// TIA Portal project "TestEssProtoFreia" (V13) (continued)

         L     #ET_MAX;
         ITD;
         DTR;
         L     #ET_MIN;
         ITD;
         DTR;
         -R;
         T     #INTER_3;  //ETENDUE DE MESURE MAXI - MINI

         L     #VAL_MINI;
         T     #INTER_4;  //ECHELLE MINI

         L     #INTER_1;
         L     #INTER_2;
         *R;
         L     #INTER_3;
         /R;
         L     #INTER_4;
         +R;
         T     #PV;
         JU    NEXT;
END_REGION

REGION Network 3 (STL): Input type : PT100 en °C
   // Input type : PT100 en °C

   C2:   L     #INPUT;
         ITD;
         DTR;
         L     10.0;
         /R;
         T     #INTER_1;



         L     #INTER_1;
         T     #PV;

         JU    NEXT;
END_REGION

REGION Network 4 (STL): Input type : PT100 en K
   // Input type  : PT100 en K

   C3:   L     #INPUT;
         ITD;
         DTR;
         L     10.0;
         /R;
         L     273.0;
         +R;
         T     #INTER_1;



         L     #INTER_1;
         T     #PV;

         JU    NEXT;
END_REGION

REGION Network 5 (STL): Depassement haut de la valeur convertie
   // Dépassement haut et bas process de la valeur
   NEXT: L     #PV;
         L     #PV_SEUILH;  //Test la valeur maximum pour le dépassement haut
         >R;
         =     #ALM_HIGH;

         L     #PV;
         L     #PV_SEUILB;  //Test la valeur minimum pour le dépassement bas
         <R;
         =     #ALM_LOW;
END_REGION

REGION Network 6 (STL): Depassement bas de la valeur convertie
   // Défaut capteur

         L     #INPUT;
         L     #ET_MAX;
         >I;
         O(;
         L     #INPUT;
         L     #ET_MIN;
         <I;
         );
         =     #ALM_TEMP;

         A     #ALM_TEMP;
         S     #ALM_SENSOR;

         AN    #ALM_TEMP;
         A     #ACQ;
         R     #ALM_SENSOR;

         NOP   0;
END_REGION

REGION Network 7 (STL): Recopie des mini et maxi de la mesure
   // Recopie des mini et maxi de la mesure
         L     #VAL_MAXI;  //Charge le maxi
         T     #PV_HIGH;

         L     #VAL_MINI;  //Charge le mini
         T     #PV_LOW;
END_REGION

REGION Network 8 (STL): Gestion du mot de défaut
   // Gestion du mot de défaut
         A     #ALM_SENSOR;
         JCN   High;  //Retourne un défaut capteur dans le mot
         L     3;  //Usually 3
         T     #ANIM;
         JU    Saut;
   High: A     #ALM_HIGH;
         JCN   Low;  //Retourne un dépassement haut dans le mot
         L     2;
         T     #ANIM;
         JU    Saut;
   Low:  A     #ALM_LOW;
         JCN   Fin;  //Retourne un dépassement bas dans le mot
         L     1;  //Usually 3
         T     #ANIM;
         JU    Saut;

   Fin:  L     0;  //Aucun défaut sur la mesure
         T     #ANIM;
   Saut: NOP   0;
END_REGION

REGION Network 9 (STL): Fin du traitement
   // Fin du traitement
   End:  NOP   0;
END_REGION
END_FUNCTION

FUNCTION "CONVERSION R/T" : Void   // FC20, SCL
{ S7_Optimized_Access := 'FALSE' }
VERSION : 0.1
BEGIN

   //#TEMPERATURE_KELVIN := REAL#29.377125832 + (REAL#2.3156100732 * #"RESISTANCE _OHMS") + (REAL#1.2102319168 * 10 ** -03 * SQR(#"RESISTANCE _OHMS"));
   #TEMPERATURE_KELVIN := REAL#29.37713 + (REAL#2.315610 * #"RESISTANCE _OHMS") + (REAL#1.210232 * 10 ** -03 * SQR(#"RESISTANCE _OHMS"));
END_FUNCTION

FUNCTION "Send_to_Epics" : Void   // FC30, LAD
{ S7_Optimized_Access := 'FALSE' }
VERSION : 0.1
   VAR_TEMP   // added for the SCL form of the ladder/FBD networks
      _w1 : Bool;
   END_VAR
BEGIN

REGION Network 1 (STL): Send timer
         AN    "EPICS_send_T1";
         L     s5t#100ms;
         SD    "EPICS_send_T0";
         A     "EPICS_send_T0";
         L     s5t#100ms;
         SD    "EPICS_send_T1";
         =     "EPICS_do_send";
END_REGION

REGION Network 2: Set ACT_SEND
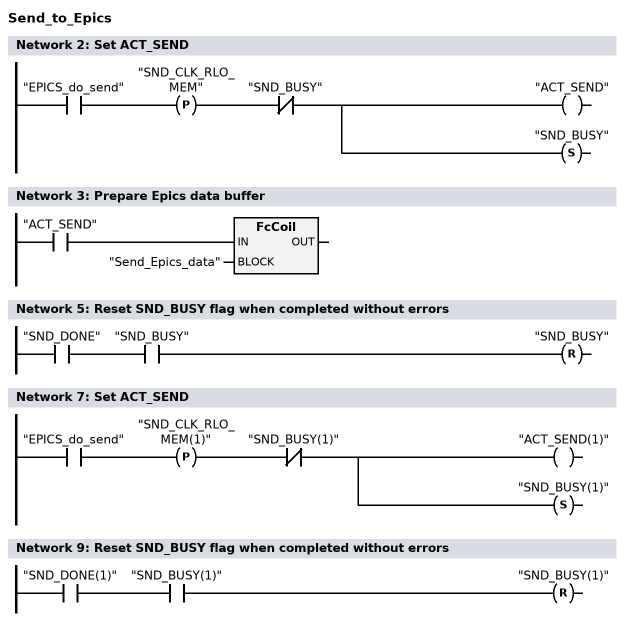
   RUNG wire#powerrail
      Contact( "EPICS_do_send" )
      P_Trig( "SND_CLK_RLO_MEM" )
      I_Contact( "SND_BUSY" )
      wire#w1
      Coil( "ACT_SEND" )
   END_RUNG
   RUNG wire#w1
      S_Coil( "SND_BUSY" )
   END_RUNG
   // the same network as SCL:
   #_w1 := "EPICS_do_send" AND NOT "SND_CLK_RLO_MEM";   // rising edge
   "SND_CLK_RLO_MEM" := "EPICS_do_send";
   "ACT_SEND" := #_w1 AND NOT "SND_BUSY";
   IF "ACT_SEND" THEN "SND_BUSY" := TRUE; END_IF;
END_REGION

REGION Network 3: Prepare Epics data buffer
   // no SCL statement known for FcCoil: written as a call
   FcCoil(block := "Send_Epics_data", in := "ACT_SEND");
END_REGION

REGION Network 4 (STL): Call AG_SEND
         CALL  AG_SEND
         ( ACT    := "ACT_SEND",
           ID     := 1,
           LADDR  := w#16#400,
           SEND   := P#DB100.DBX0.0 BYTE 2000,
           LEN    := 2000,
           DONE   := "SND_DONE",
           ERROR  := "SND_ERR",
           STATUS := "SEND_status"
         );
END_REGION

REGION Network 5: Reset SND_BUSY flag when completed without errors
   RUNG wire#powerrail
      Contact( "SND_DONE" )
      Contact( "SND_BUSY" )
      R_Coil( "SND_BUSY" )
   END_RUNG
   // the same network as SCL:
   IF "SND_DONE" AND "SND_BUSY" THEN "SND_BUSY" := FALSE; END_IF;
END_REGION

REGION Network 6 (STL): Reset SND_BUSY flag and save the status when returned error
         AN    "SND_DONE";
         A     "SND_ERR";
         JNB   ex1;
         R     "SND_BUSY";
         L     "SEND_status";
         T     "SND_STAT_SAVE";
   ex1:  NOP   0;
END_REGION

REGION Network 7: Set ACT_SEND
   RUNG wire#powerrail
      Contact( "EPICS_do_send" )
      P_Trig( "SND_CLK_RLO_MEM(1)" )
      I_Contact( "SND_BUSY(1)" )
      wire#w1
      Coil( "ACT_SEND(1)" )
   END_RUNG
   RUNG wire#w1
      S_Coil( "SND_BUSY(1)" )
   END_RUNG
   // the same network as SCL:
   #_w1 := "EPICS_do_send" AND NOT "SND_CLK_RLO_MEM(1)";   // rising edge
   "SND_CLK_RLO_MEM(1)" := "EPICS_do_send";
   "ACT_SEND(1)" := #_w1 AND NOT "SND_BUSY(1)";
   IF "ACT_SEND(1)" THEN "SND_BUSY(1)" := TRUE; END_IF;
END_REGION

REGION Network 8 (STL): Call AG_SEND
         CALL  AG_SEND
         ( ACT    := "ACT_SEND(1)",
           ID     := 2,
           LADDR  := w#16#400,
           SEND   := P#DB104.DBX0.0 BYTE 40,
           LEN    := 40,
           DONE   := "SND_DONE(1)",
           ERROR  := "SND_ERR(1)",
           STATUS := "SEND_status(1)"
         );
END_REGION

REGION Network 9: Reset SND_BUSY flag when completed without errors
   RUNG wire#powerrail
      Contact( "SND_DONE(1)" )
      Contact( "SND_BUSY(1)" )
      R_Coil( "SND_BUSY(1)" )
   END_RUNG
   // the same network as SCL:
   IF "SND_DONE(1)" AND "SND_BUSY(1)" THEN "SND_BUSY(1)" := FALSE; END_IF;
END_REGION

REGION Network 10 (STL): Reset SND_BUSY flag and save the status when returned error
         AN    "SND_DONE(1)";
         A     "SND_ERR(1)";
         JNB   ex2;
         R     "SND_BUSY(1)";
         L     "SEND_status(1)";
         T     "SND_STAT_SAVE(1)";
   ex2:  NOP   0;
END_REGION
END_FUNCTION

FUNCTION "Recv_from_Epics" : Void   // FC31, STL
{ S7_Optimized_Access := 'FALSE' }
VERSION : 0.1
BEGIN

REGION Network 1: Get data from Epics (channel 1)
         CALL  AG_RECV
         ( ID     := 1,
           LADDR  := w#16#400,
           RECV   := P#DB101.DBX0.0 BYTE 1000,
           NDR    := "RCV_NDR",
           ERROR  := "RCV_ERR",
           STATUS := "RECV_status",
           LEN    := "RECV_len"
         );
         AN    "RCV_NDR";
         O     "RCV_ERR";
         JC    out;
         CALL  "Cmds_from_Epics";
         BE;
   out:  AN    "RCV_ERR";
         JC    _001;
         L     "RECV_status";
         T     "RCV_STAT_SAVE";
   _001: NOP   0;
END_REGION

REGION Network 2: Get data from Epics (channel 2)
         CALL  AG_RECV
         ( ID     := 2,
           LADDR  := w#16#400,
           RECV   := P#DB105.DBX0.0 BYTE 250,
           NDR    := "RCV_NDR(1)",
           ERROR  := "RCV_ERR(1)",
           STATUS := "RECV_status(1)",
           LEN    := "RECV_len(1)"
         );
         AN    "RCV_NDR(1)";
         O     "RCV_ERR(1)";
         JC    out2;
         CALL  "Data_from_IOC";
         BE;
   out2: AN    "RCV_ERR(1)";
         JC    _002;
         L     "RECV_status(1)";
         T     "RCV_STAT_SAVE(1)";
   _002: NOP   0;
END_REGION
END_FUNCTION

FUNCTION "Send_Epics_data" : Void   // FC32, STL
{ S7_Optimized_Access := 'FALSE' }
VERSION : 0.1
BEGIN

REGION Network 2: Update the Local/remote status
         A     "LocalMode";
         =     "PLC_to_Epics".sLocal;
END_REGION

REGION Network 3: CV01
         L     "CV01_HMI_VAL";
         T     "PLC_to_Epics".CV01.sSetV;
         L     "Tag_7";
         T     "PLC_to_Epics".CV01.sRdV;

         AN    "CV01_ManAuto";
         =     "PLC_to_Epics".CV01.sAuto;
END_REGION

REGION Network 4: CV02
         L     "CV02_HMI_VAL";
         T     "PLC_to_Epics".CV02.sSetV;
         L     "Tag_8";
         T     "PLC_to_Epics".CV02.sRdV;

         AN    "CV02_ManAuto";
         =     "PLC_to_Epics".CV02.sAuto;
END_REGION

REGION Network 5: CV03
         L     "CV03_HMI_VAL";
         T     "PLC_to_Epics".CV03.sSetV;
         L     "Tag_9";
         T     "PLC_to_Epics".CV03.sRdV;

         AN    "CV03_ManAuto";
         =     "PLC_to_Epics".CV03.sAuto;
END_REGION

REGION Network 6: CV04
         L     "CV04_HMI_VAL";
         T     "PLC_to_Epics".CV04.sSetV;
         L     "Tag_10";
         T     "PLC_to_Epics".CV04.sRdV;

         AN    "CV04_ManAuto";
         =     "PLC_to_Epics".CV04.sAuto;
END_REGION

REGION Network 7: CV05
         L     "CV05_HMI_VAL";
         T     "PLC_to_Epics".CV05.sSetV;
         L     "Tag_11";
         T     "PLC_to_Epics".CV05.sRdV;

   //      AN    "CV05_ManAuto"
   //      =     "PLC_to_Epics".CV05.sAuto
END_REGION

REGION Network 8: CV07
         L     "CV07_HMI_VAL";
         T     "PLC_to_Epics".CV07.sSetV;
         L     "Tag_12";
         T     "PLC_to_Epics".CV07.sRdV;

         AN    "CV07_ManAuto";
         =     "PLC_to_Epics".CV07.sAuto;
END_REGION

REGION Network 9: CV60
         L     "CV60_HMI_VAL";
         T     "PLC_to_Epics".CV60.sSetV;
         L     "Tag_13";
         T     "PLC_to_Epics".CV60.sRdV;

         AN    "CV60_ManAuto";
         =     "PLC_to_Epics".CV60.sAuto;
END_REGION

REGION Network 10: CV61
         L     "CV61_HMI_VAL";
         T     "PLC_to_Epics".CV61.sSetV;
         L     "Tag_14";
         T     "PLC_to_Epics".CV61.sRdV;

         AN    "CV61_ManAuto";
         =     "PLC_to_Epics".CV61.sAuto;
END_REGION

REGION Network 11: CV62
         L     "CV62_HMI_VAL";
         T     "PLC_to_Epics".CV62.sSetV;
         L     "Tag_15";
         T     "PLC_to_Epics".CV62.sRdV;

   //      AN    "CV62_ManAuto"
   //      =     "PLC_to_Epics".CV62.sAuto
END_REGION

REGION Network 12: CV550
         AN    "ASCOenManuel";
         =     "PLC_to_Epics".CV550.sAuto;
         =     "Data_to_HNOSS".RegOnMKS2;
END_REGION

REGION Network 13: CV550
         L     "S6_parameters".CV550;
         T     "PLC_to_Epics".CV550.sSetV;
END_REGION

REGION Network 14: spare - VB chan 7
         A     "voie 7 chaufferette BV";
         =     "PLC_to_Epics"."spare-VB-7".sHtrOn;
END_REGION

REGION Network 15: spare - VB chan 8
         A     "voie 8 chaufferette BV";
         =     "PLC_to_Epics"."spare-VB-8".sHtrOn;
END_REGION

REGION Network 16: spare VB chan 9
         A     "voie 9 chaufferette BV";
         =     "PLC_to_Epics"."spare-VB-9".sHtrOn;
END_REGION

REGION Network 17: spare - VB chan 10
         A     "voie 10  chaufferette BV";
         =     "PLC_to_Epics"."spare-VB-10".sHtrOn;
END_REGION

REGION Network 18: spare - VB chan 11
         A     "voie 11 chaufferette BV";
         =     "PLC_to_Epics"."spare-VB-11".sHtrOn;
END_REGION

REGION Network 19: spare - CM chan 5
         A     "voie 5 chaufferette CM";
         =     "PLC_to_Epics"."spare-CM-5".sHtrOn;
END_REGION

REGION Network 20: spare - CM chan 6
         A     "voie 6 chaufferette CM";
         =     "PLC_to_Epics"."spare-CM-6".sHtrOn;
END_REGION

REGION Network 21: spare - CM chan 7
         A     "voie 7 chaufferette CM";
         =     "PLC_to_Epics"."spare-CM-7".sHtrOn;
END_REGION

REGION Network 22: spare - CM chan 8
         A     "voie 8 chaufferette CM";
         =     "PLC_to_Epics"."spare-CM-8".sHtrOn;
END_REGION

REGION Network 23: spare - CM chan 10
         A     "voie 10 chaufferette CM";
         =     "PLC_to_Epics"."spare-CM-10".sHtrOn;
END_REGION

REGION Network 24: spare - CM chan 12
         A     "voie 12 chaufferette CM";
         =     "PLC_to_Epics"."spare-CM-12".sHtrOn;
END_REGION

REGION Network 25: Status bits
         A     "Graph/manuelle";
         =     "PLC_to_Epics".sManual;
         A     "ErreurSupervision";
         =     "PLC_to_Epics".sGrafcetERR;
         A     "Etat initial";
         =     "PLC_to_Epics".sGS1;
         A     "EtatCdtCryo";
         =     "PLC_to_Epics".sGS2;
         A     "EtatAttMef";
         =     "PLC_to_Epics".sGS3;
         A     "EtatMEFazote";
         =     "PLC_to_Epics".sGS4;
         A     "EtatMEFhelium";
         =     "PLC_to_Epics".sGS5;
         A     "EtatMode4k";
         =     "PLC_to_Epics".sGS6;
         A     "EtatModeStandBy";
         =     "PLC_to_Epics".sGS7;
         A     "EtatMode2K";
         =     "PLC_to_Epics".sGS8;
         A     "Etatrechauffage";
         =     "PLC_to_Epics".sGS10;
         A     "conditionTempMEFheliumOK";
         =     "PLC_to_Epics".sTransTempOK;
         A     "TransMode4K";
         =     "PLC_to_Epics".sTransMode4K;
         A     "EPICS_COMM_OK";
         =     "PLC_to_Epics".EpicsCommOK;
         A     "HNOSS_COMM_OK";
         =     "PLC_to_Epics".HNOSSCommOK;
END_REGION

REGION Network 26: Real parameters read-back (LHe level PID settings)
         L     "S8_parameters".TrigPID_CV01;
         T     "PLC_to_Epics".TrigPID_CV01.sSetV;
         L     "S6_parameters".TrigPID_CV02;
         T     "PLC_to_Epics".TrigPID_CV02.sSetV;
         L     "S6_parameters".TrigPID_CV03;
         T     "PLC_to_Epics".TrigPID_CV03.sSetV;
         L     "S8_parameters".PID_LT01_CV01_SP;
         T     "PLC_to_Epics".PID_LT01_CV01_SP.sSetV;
         L     "S6_parameters".PID_LT01_CV02_SP;
         T     "PLC_to_Epics".PID_LT01_CV02_SP.sSetV;
         L     "S6_parameters".PID_LT03_CV03_SP;
         T     "PLC_to_Epics".PID_LT03_CV03_SP.sSetV;
END_REGION

REGION Network 27: Real parameters read-back (CV550l PID settings)
         L     "S6_parameters".PID_PT01_CV550_SP;
         T     "PLC_to_Epics".PID_PT01_CV550_SP.sSetV;
END_REGION

REGION Network 28: Sequence steps
         L     "Data_to_HNOSS".S4step;
         T     "PLC_to_Epics".S4step;
         L     "Data_to_HNOSS".S5step;
         T     "PLC_to_Epics".S5step;
         L     "Data_to_HNOSS".S6step;
         T     "PLC_to_Epics".S6step;
         L     "Data_to_HNOSS".S7step;
         T     "PLC_to_Epics".S7step;
         L     "Data_to_HNOSS".S8step;
         T     "PLC_to_Epics".S8step;
         L     "Data_to_HNOSS".S9step;
         T     "PLC_to_Epics".S9step;
         L     "Data_to_HNOSS".S10step;
         T     "PLC_to_Epics".S10step;
         L     "Data_to_HNOSS".SXstep;
         T     "PLC_to_Epics".SXstep;
END_REGION

REGION Network 29: PID's GAINS
         L     "S8_parameters".CV01_PID_GAIN;
         T     "PLC_to_Epics".CV01_PID_GAIN.sSetV;
         L     "S6_parameters".CV02_PID_GAIN;
         T     "PLC_to_Epics".CV02_PID_GAIN.sSetV;
         L     "S6_parameters".CV03_PID_GAIN;
         T     "PLC_to_Epics".CV03_PID_GAIN.sSetV;
         L     "S4_Parameters".CV60_PID_GAIN;
         T     "PLC_to_Epics".CV60_PID_GAIN.sSetV;
END_REGION

REGION Network 30: CV01 PID TI
         A(;
         L     "S8_parameters".CV01_PID_TI;
         DTR;
         T     #tmpR;
         SET;
         SAVE;
         CLR;
         A     BR;
         );
         JNB   Label_0;
         L     #tmpR;
         L     1000.0;
         /R;
         T     "PLC_to_Epics".CV01_PID_TI.sSetV;
   Label_0:NOP   0;
END_REGION

REGION Network 31: CV01 PID TD
         A(;
         L     "S8_parameters".CV01_PID_TD;
         DTR;
         T     #tmpR;
         SET;
         SAVE;
         CLR;
         A     BR;
         );
         JNB   Label_1;
         L     #tmpR;
         L     1000.0;
         /R;
         T     "PLC_to_Epics".CV01_PID_TD.sSetV;
   Label_1:NOP   0;
END_REGION

REGION Network 32: CV01 PID TM_LAG
         A(;
         L     "S8_parameters".CV01_PID_TM_LAG;
         DTR;
         T     #tmpR;
         SET;
         SAVE;
         CLR;
         A     BR;
         );
         JNB   Label_2;
         L     #tmpR;
         L     1000.0;
         /R;
         T     "PLC_to_Epics".CV01_PID_TM_LAG.sSetV;
   Label_2:NOP   0;
END_REGION

REGION Network 33: CV02 PID TI
         A(;
         L     "S6_parameters".CV02_PID_TI;
         DTR;
         T     #tmpR;
         SET;
         SAVE;
         CLR;
         A     BR;
         );
         JNB   Label_3;
         L     #tmpR;
         L     1000.0;
         /R;
         T     "PLC_to_Epics".CV02_PID_TI.sSetV;
   Label_3:NOP   0;
END_REGION

REGION Network 34: CV02 PID TD
         A(;
         L     "S6_parameters".CV02_PID_TD;
         DTR;
         T     #tmpR;
         SET;
         SAVE;
         CLR;
         A     BR;
         );
         JNB   Label_4;
         L     #tmpR;
         L     1000.0;
         /R;
         T     "PLC_to_Epics".CV02_PID_TD.sSetV;
   Label_4:NOP   0;
END_REGION

REGION Network 35: CV02 PID TM_LAG
         A(;
         L     "S6_parameters".CV02_PID_TM_LAG;
         DTR;
         T     #tmpR;
         SET;
         SAVE;
         CLR;
         A     BR;
         );
         JNB   Label_5;
         L     #tmpR;
         L     1000.0;
         /R;
         T     "PLC_to_Epics".CV02_PID_TM_LAG.sSetV;
   Label_5:NOP   0;
END_REGION

REGION Network 36: CV03 PID TI
         A(;
         L     "S6_parameters".CV03_PID_TI;
         DTR;
         T     #tmpR;
         SET;
         SAVE;
         CLR;
         A     BR;
         );
         JNB   Label_6;
         L     #tmpR;
         L     1000.0;
         /R;
         T     "PLC_to_Epics".CV03_PID_TI.sSetV;
   Label_6:NOP   0;
END_REGION

REGION Network 37: CV03 PID TD
         A(;
         L     "S6_parameters".CV03_PID_TD;
         DTR;
         T     #tmpR;
         SET;
         SAVE;
         CLR;
         A     BR;
         );
         JNB   Label_7;
         L     #tmpR;
         L     1000.0;
         /R;
         T     "PLC_to_Epics".CV03_PID_TD.sSetV;
   Label_7:NOP   0;
END_REGION

REGION Network 38: CV03 PID TM_LAG
         A(;
         L     "S6_parameters".CV03_PID_TM_LAG;
         DTR;
         T     #tmpR;
         SET;
         SAVE;
         CLR;
         A     BR;
         );
         JNB   Label_8;
         L     #tmpR;
         L     1000.0;
         /R;
         T     "PLC_to_Epics".CV03_PID_TM_LAG.sSetV;
   Label_8:NOP   0;
END_REGION

REGION Network 39: CV60 PID TI
         A(;
         L     "S4_Parameters".CV60_PID_TI;
         DTR;
         T     #tmpR;
         SET;
         SAVE;
         CLR;
         A     BR;
         );
         JNB   Label_9;
         L     #tmpR;
         L     1000.0;
         /R;
         T     "PLC_to_Epics".CV60_PID_TI.sSetV;
   Label_9:NOP   0;
END_REGION

REGION Network 40: CV60 PID TD
         A(;
         L     "S4_Parameters".CV60_PID_TD;
         DTR;
         T     #tmpR;
         SET;
         SAVE;
         CLR;
         A     BR;
         );
         JNB   Label_10;
         L     #tmpR;
         L     1000.0;
         /R;
         T     "PLC_to_Epics".CV60_PID_TD.sSetV;
   Label_10:NOP   0;
END_REGION

REGION Network 41: CV60 PID TM_LAG
         A(;
         L     "S4_Parameters".CV60_PID_TM_LAG;
         DTR;
         T     #tmpR;
         SET;
         SAVE;
         CLR;
         A     BR;
         );
         JNB   Label_11;
         L     #tmpR;
         L     1000.0;
         /R;
         T     "PLC_to_Epics".CV60_PID_TM_LAG.sSetV;
   Label_11:NOP   0;
END_REGION

REGION Network 42: TT77_CV60 SP
         L     "S4_Parameters".CV60_PID_SP_INT;
         T     "PLC_to_Epics".PID_TT77_CV60_SP.sSetV;
END_REGION

REGION Network 43: S5/S6 parameters
         L     "S6_parameters".S5_P_FT552_MIN_GB;
         T     "PLC_to_Epics".S5_P_FT552_MIN_GB.sSetV;
         L     "S6_parameters".S5_P_FT552_MIN_C;
         T     "PLC_to_Epics".S5_P_FT552_MIN_C.sSetV;
         L     "S6_parameters".S5_P_FT552_MAX_GB;
         T     "PLC_to_Epics".S5_P_FT552_MAX_GB.sSetV;
         L     "S6_parameters".S5_P_FT552_MAX_C;
         T     "PLC_to_Epics".S5_P_FT552_MAX_C.sSetV;
END_REGION

REGION Network 44: S8_P_CV01 and S8_P_CV01_Step7
         L     "S8_parameters".S8_P_CV01;
         T     "PLC_to_Epics".S8_P_CV01.sSetV;
         L     "S8_parameters".S8_P_CV01_Step7;
         T     "PLC_to_Epics".S8_P_CV01_Step7.sSetV;
END_REGION
END_FUNCTION

FUNCTION "Cmds_from_Epics" : Void   // FC33, LAD
TITLE = Process data from Epics
{ S7_Optimized_Access := 'FALSE' }
VERSION : 0.1
   VAR_TEMP   // added for the SCL form of the ladder/FBD networks
      _w1 : Bool;
   END_VAR
BEGIN

REGION Network 1: Switch to remote mode (control from Epics)
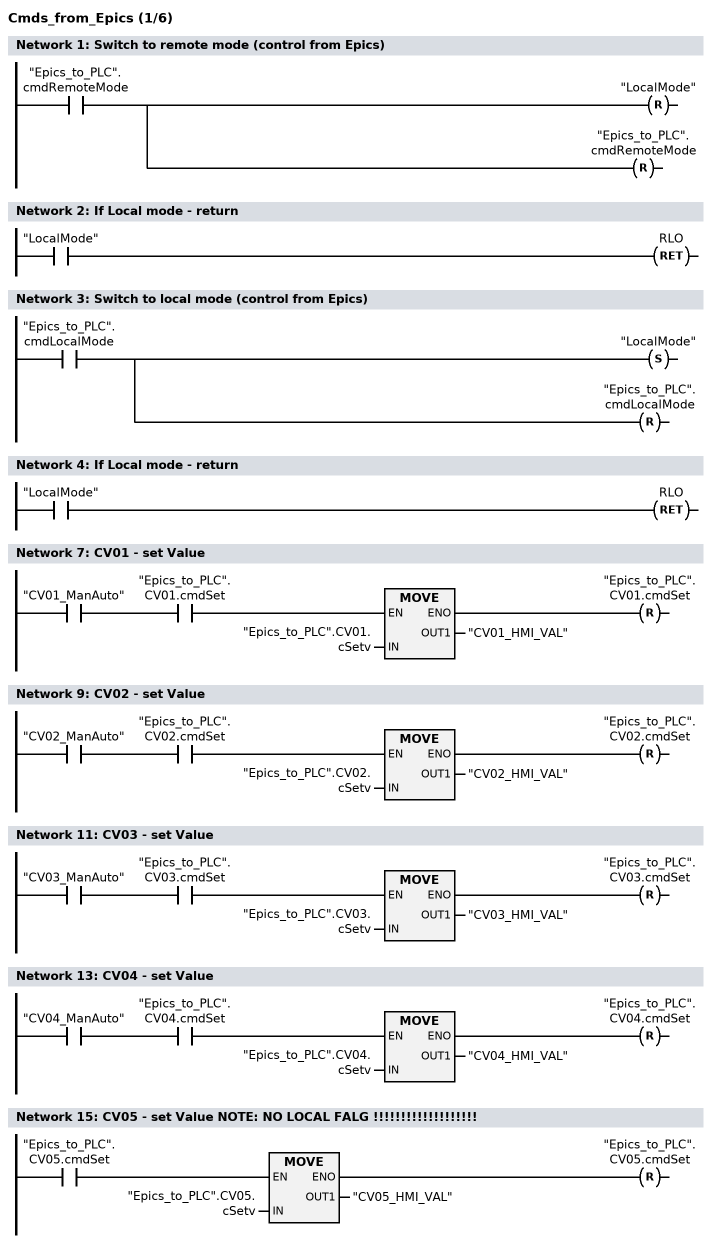
   RUNG wire#powerrail
      Contact( "Epics_to_PLC".cmdRemoteMode )
      wire#w1
      R_Coil( "LocalMode" )
   END_RUNG
   RUNG wire#w1
      R_Coil( "Epics_to_PLC".cmdRemoteMode )
   END_RUNG
   // the same network as SCL:
   IF "Epics_to_PLC".cmdRemoteMode THEN
       "LocalMode" := FALSE;
       "Epics_to_PLC".cmdRemoteMode := FALSE;
   END_IF;
END_REGION

REGION Network 2: If Local mode - return
   IF "LocalMode" THEN
       ENO := TRUE;
       RETURN;
   END_IF;
END_REGION

REGION Network 3: Switch to local mode (control from Epics)
   RUNG wire#powerrail
      Contact( "Epics_to_PLC".cmdLocalMode )
      wire#w1
      S_Coil( "LocalMode" )
   END_RUNG
   RUNG wire#w1
      R_Coil( "Epics_to_PLC".cmdLocalMode )
   END_RUNG
   // the same network as SCL:
   IF "Epics_to_PLC".cmdLocalMode THEN
       "LocalMode" := TRUE;
       "Epics_to_PLC".cmdLocalMode := FALSE;
   END_IF;
END_REGION

REGION Network 4: If Local mode - return
   IF "LocalMode" THEN
       ENO := TRUE;
       RETURN;
   END_IF;
END_REGION

REGION Network 5: Test data (copy block of data)
END_REGION

REGION Network 6 (STL): CV01 Man/Auto
         A     "Epics_to_PLC".CV01.cmdAuto;
         R     "CV01_ManAuto";
         A     "Epics_to_PLC".CV01.cmdMan;
         S     "CV01_ManAuto";
END_REGION

REGION Network 7: CV01 - set Value
   RUNG wire#powerrail
      Contact( "CV01_ManAuto" )
      Contact( "Epics_to_PLC".CV01.cmdSet )
      { S7_GenerateENO := "TRUE" } Move(in := "Epics_to_PLC".CV01.cSetv, out1 => "CV01_HMI_VAL")
      R_Coil( "Epics_to_PLC".CV01.cmdSet )
   END_RUNG
   // the same network as SCL:
   // ENO of a box is taken as its EN; it also drops when the box reports an error
   IF "CV01_ManAuto" AND "Epics_to_PLC".CV01.cmdSet THEN
       "CV01_HMI_VAL" := "Epics_to_PLC".CV01.cSetv;
       "Epics_to_PLC".CV01.cmdSet := FALSE;
   END_IF;
END_REGION

REGION Network 8 (STL): CV02 Man/Auto
         A     "Epics_to_PLC".CV02.cmdAuto;
         R     "CV02_ManAuto";
         A     "Epics_to_PLC".CV02.cmdMan;
         S     "CV02_ManAuto";
END_REGION

REGION Network 9: CV02 - set Value
   RUNG wire#powerrail
      Contact( "CV02_ManAuto" )
      Contact( "Epics_to_PLC".CV02.cmdSet )
      { S7_GenerateENO := "TRUE" } Move(in := "Epics_to_PLC".CV02.cSetv, out1 => "CV02_HMI_VAL")
      R_Coil( "Epics_to_PLC".CV02.cmdSet )
   END_RUNG
   // the same network as SCL:
   // ENO of a box is taken as its EN; it also drops when the box reports an error
   IF "CV02_ManAuto" AND "Epics_to_PLC".CV02.cmdSet THEN
       "CV02_HMI_VAL" := "Epics_to_PLC".CV02.cSetv;
       "Epics_to_PLC".CV02.cmdSet := FALSE;
   END_IF;
END_REGION

REGION Network 10 (STL): CV03 Man/Auto
         A     "Epics_to_PLC".CV03.cmdAuto;
         R     "CV03_ManAuto";
         A     "Epics_to_PLC".CV03.cmdMan;
         S     "CV03_ManAuto";
END_REGION

REGION Network 11: CV03 - set Value
   RUNG wire#powerrail
      Contact( "CV03_ManAuto" )
      Contact( "Epics_to_PLC".CV03.cmdSet )
      { S7_GenerateENO := "TRUE" } Move(in := "Epics_to_PLC".CV03.cSetv, out1 => "CV03_HMI_VAL")
      R_Coil( "Epics_to_PLC".CV03.cmdSet )
   END_RUNG
   // the same network as SCL:
   // ENO of a box is taken as its EN; it also drops when the box reports an error
   IF "CV03_ManAuto" AND "Epics_to_PLC".CV03.cmdSet THEN
       "CV03_HMI_VAL" := "Epics_to_PLC".CV03.cSetv;
       "Epics_to_PLC".CV03.cmdSet := FALSE;
   END_IF;
END_REGION

REGION Network 12 (STL): CV04 Man/Auto
         A     "Epics_to_PLC".CV04.cmdAuto;
         R     "CV04_ManAuto";
         A     "Epics_to_PLC".CV04.cmdMan;
         S     "CV04_ManAuto";
END_REGION

REGION Network 13: CV04 - set Value
   RUNG wire#powerrail
      Contact( "CV04_ManAuto" )
      Contact( "Epics_to_PLC".CV04.cmdSet )
      { S7_GenerateENO := "TRUE" } Move(in := "Epics_to_PLC".CV04.cSetv, out1 => "CV04_HMI_VAL")
      R_Coil( "Epics_to_PLC".CV04.cmdSet )
   END_RUNG
   // the same network as SCL:
   // ENO of a box is taken as its EN; it also drops when the box reports an error
   IF "CV04_ManAuto" AND "Epics_to_PLC".CV04.cmdSet THEN
       "CV04_HMI_VAL" := "Epics_to_PLC".CV04.cSetv;
       "Epics_to_PLC".CV04.cmdSet := FALSE;
   END_IF;
END_REGION

REGION Network 14: CV05 Man/Auto
END_REGION

REGION Network 15: CV05 - set Value NOTE: NO LOCAL FALG !!!!!!!!!!!!!!!!!!!
   RUNG wire#powerrail
      Contact( "Epics_to_PLC".CV05.cmdSet )
      { S7_GenerateENO := "TRUE" } Move(in := "Epics_to_PLC".CV05.cSetv, out1 => "CV05_HMI_VAL")
      R_Coil( "Epics_to_PLC".CV05.cmdSet )
   END_RUNG
   // the same network as SCL:
   // ENO of a box is taken as its EN; it also drops when the box reports an error
   IF "Epics_to_PLC".CV05.cmdSet THEN
       "CV05_HMI_VAL" := "Epics_to_PLC".CV05.cSetv;
       "Epics_to_PLC".CV05.cmdSet := FALSE;
   END_IF;
END_REGION

REGION Network 16 (STL): CV07 Man/Auto
         A     "Epics_to_PLC".CV07.cmdAuto;
         R     "CV07_ManAuto";
         A     "Epics_to_PLC".CV07.cmdMan;
         S     "CV07_ManAuto";
END_REGION

REGION Network 17: CV07 - set Value
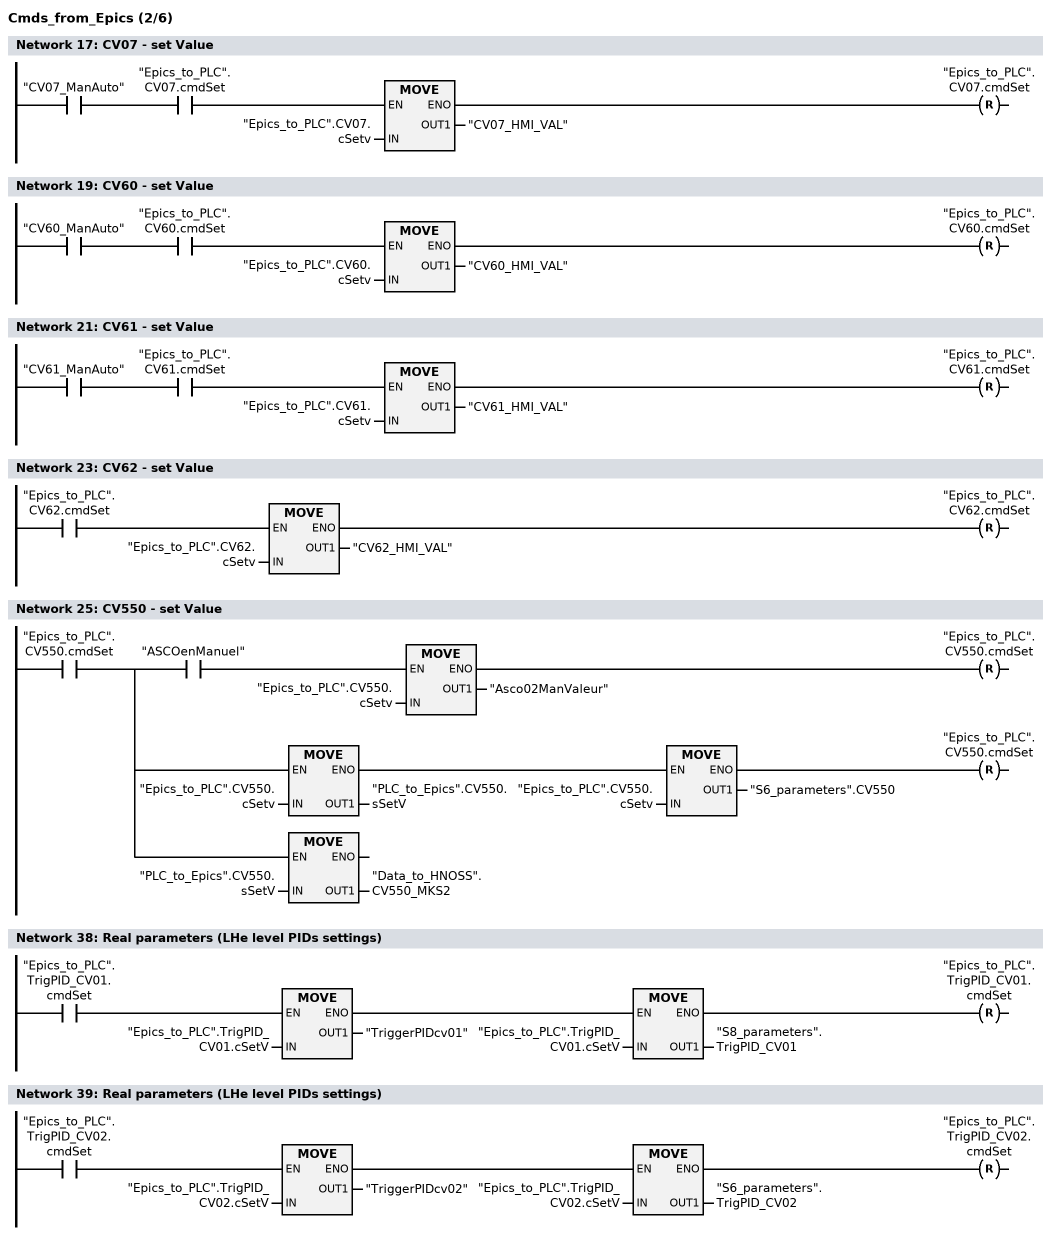
   RUNG wire#powerrail
      Contact( "CV07_ManAuto" )
      Contact( "Epics_to_PLC".CV07.cmdSet )
      { S7_GenerateENO := "TRUE" } Move(in := "Epics_to_PLC".CV07.cSetv, out1 => "CV07_HMI_VAL")
      R_Coil( "Epics_to_PLC".CV07.cmdSet )
   END_RUNG
   // the same network as SCL:
   // ENO of a box is taken as its EN; it also drops when the box reports an error
   IF "CV07_ManAuto" AND "Epics_to_PLC".CV07.cmdSet THEN
       "CV07_HMI_VAL" := "Epics_to_PLC".CV07.cSetv;
       "Epics_to_PLC".CV07.cmdSet := FALSE;
   END_IF;
END_REGION

REGION Network 18 (STL): CV60 Man/Auto
         A     "Epics_to_PLC".CV60.cmdAuto;
         R     "CV60_ManAuto";
         A     "Epics_to_PLC".CV60.cmdMan;
         S     "CV60_ManAuto";
END_REGION

REGION Network 19: CV60 - set Value
   RUNG wire#powerrail
      Contact( "CV60_ManAuto" )
      Contact( "Epics_to_PLC".CV60.cmdSet )
      { S7_GenerateENO := "TRUE" } Move(in := "Epics_to_PLC".CV60.cSetv, out1 => "CV60_HMI_VAL")
      R_Coil( "Epics_to_PLC".CV60.cmdSet )
   END_RUNG
   // the same network as SCL:
   // ENO of a box is taken as its EN; it also drops when the box reports an error
   IF "CV60_ManAuto" AND "Epics_to_PLC".CV60.cmdSet THEN
       "CV60_HMI_VAL" := "Epics_to_PLC".CV60.cSetv;
       "Epics_to_PLC".CV60.cmdSet := FALSE;
   END_IF;
END_REGION

REGION Network 20 (STL): CV61 Man/Auto
         A     "Epics_to_PLC".CV61.cmdAuto;
         R     "CV61_ManAuto";
         A     "Epics_to_PLC".CV61.cmdMan;
         S     "CV61_ManAuto";
END_REGION

REGION Network 21: CV61 - set Value
   RUNG wire#powerrail
      Contact( "CV61_ManAuto" )
      Contact( "Epics_to_PLC".CV61.cmdSet )
      { S7_GenerateENO := "TRUE" } Move(in := "Epics_to_PLC".CV61.cSetv, out1 => "CV61_HMI_VAL")
      R_Coil( "Epics_to_PLC".CV61.cmdSet )
   END_RUNG
   // the same network as SCL:
   // ENO of a box is taken as its EN; it also drops when the box reports an error
   IF "CV61_ManAuto" AND "Epics_to_PLC".CV61.cmdSet THEN
       "CV61_HMI_VAL" := "Epics_to_PLC".CV61.cSetv;
       "Epics_to_PLC".CV61.cmdSet := FALSE;
   END_IF;
END_REGION

REGION Network 22: CV62 Man/Auto
END_REGION

REGION Network 23: CV62 - set Value
   RUNG wire#powerrail
      Contact( "Epics_to_PLC".CV62.cmdSet )
      { S7_GenerateENO := "TRUE" } Move(in := "Epics_to_PLC".CV62.cSetv, out1 => "CV62_HMI_VAL")
      R_Coil( "Epics_to_PLC".CV62.cmdSet )
   END_RUNG
   // the same network as SCL:
   // ENO of a box is taken as its EN; it also drops when the box reports an error
   IF "Epics_to_PLC".CV62.cmdSet THEN
       "CV62_HMI_VAL" := "Epics_to_PLC".CV62.cSetv;
       "Epics_to_PLC".CV62.cmdSet := FALSE;
   END_IF;
END_REGION

REGION Network 24 (STL): CV550 Man/Auto
         A     "Epics_to_PLC".CV550.cmdAuto;
         R     "ASCOenManuel";
         A     "Epics_to_PLC".CV550.cmdMan;
         S     "ASCOenManuel";
END_REGION

REGION Network 25: CV550 - set Value
   RUNG wire#powerrail
      Contact( "Epics_to_PLC".CV550.cmdSet )
      wire#w1
      Contact( "ASCOenManuel" )
      { S7_GenerateENO := "TRUE" } Move(in := "Epics_to_PLC".CV550.cSetv, out1 => "Asco02ManValeur")
      R_Coil( "Epics_to_PLC".CV550.cmdSet )
   END_RUNG
   RUNG wire#w1
      { S7_GenerateENO := "TRUE" } Move(in := "Epics_to_PLC".CV550.cSetv, out1 => "PLC_to_Epics".CV550.sSetV)
      { S7_GenerateENO := "TRUE" } Move(in := "Epics_to_PLC".CV550.cSetv, out1 => "S6_parameters".CV550)
      R_Coil( "Epics_to_PLC".CV550.cmdSet )
   END_RUNG
   RUNG wire#w1
      { S7_GenerateENO := "TRUE" } Move(in := "PLC_to_Epics".CV550.sSetV, out1 => "Data_to_HNOSS".CV550_MKS2)
   END_RUNG
   // the same network as SCL:
   // ENO of a box is taken as its EN; it also drops when the box reports an error
   IF "Epics_to_PLC".CV550.cmdSet AND "ASCOenManuel" THEN
       "Asco02ManValeur" := "Epics_to_PLC".CV550.cSetv;
   END_IF;
   #_w1 := "Epics_to_PLC".CV550.cmdSet;
   IF "Epics_to_PLC".CV550.cmdSet AND "ASCOenManuel" THEN "Epics_to_PLC".CV550.cmdSet := FALSE; END_IF;
   IF #_w1 THEN
       "PLC_to_Epics".CV550.sSetV := "Epics_to_PLC".CV550.cSetv;
       "S6_parameters".CV550 := "Epics_to_PLC".CV550.cSetv;
       "Epics_to_PLC".CV550.cmdSet := FALSE;
       "Data_to_HNOSS".CV550_MKS2 := "PLC_to_Epics".CV550.sSetV;
   END_IF;
END_REGION

REGION Network 26 (STL): spare- VB chan 7
         A     "Epics_to_PLC"."spare-VB-7".cmdSet;
         S     "voie 7 chaufferette BV";
         A     "Epics_to_PLC"."spare-VB-7".cmdRst;
         R     "voie 7 chaufferette BV";
END_REGION

REGION Network 27 (STL): spare- VB chan 8
         A     "Epics_to_PLC"."spare-VB-8".cmdSet;
         S     "voie 8 chaufferette BV";
         A     "Epics_to_PLC"."spare-VB-8".cmdRst;
         R     "voie 8 chaufferette BV";
END_REGION

REGION Network 28 (STL): spare- VB chan 9
         A     "Epics_to_PLC"."spare-VB-9".cmdSet;
         S     "voie 9 chaufferette BV";
         A     "Epics_to_PLC"."spare-VB-9".cmdRst;
         R     "voie 9 chaufferette BV";
END_REGION

REGION Network 29 (STL): spare- VB chan 10
         A     "Epics_to_PLC"."spare-VB-10".cmdSet;
         S     "voie 10  chaufferette BV";
         A     "Epics_to_PLC"."spare-VB-10".cmdRst;
         R     "voie 10  chaufferette BV";
END_REGION

REGION Network 30 (STL): spare - VB chan 11
         A     "Epics_to_PLC"."spare-VB-11".cmdSet;
         S     "voie 11 chaufferette BV";
         A     "Epics_to_PLC"."spare-VB-11".cmdRst;
         R     "voie 11 chaufferette BV";
END_REGION

REGION Network 31 (STL): spare - CM chan 5
         A     "Epics_to_PLC"."spare-CM-5".cmdSet;
         S     "voie 5 chaufferette CM";
         A     "Epics_to_PLC"."spare-CM-5".cmdRst;
         R     "voie 5 chaufferette CM";
END_REGION

REGION Network 32 (STL): spare - CM chan 6
         A     "Epics_to_PLC"."spare-CM-6".cmdSet;
         S     "voie 6 chaufferette CM";
         A     "Epics_to_PLC"."spare-CM-6".cmdRst;
         R     "voie 6 chaufferette CM";
END_REGION

REGION Network 33 (STL): spare - CM chan 7
         A     "Epics_to_PLC"."spare-CM-7".cmdSet;
         S     "voie 7 chaufferette CM";
         A     "Epics_to_PLC"."spare-CM-7".cmdRst;
         R     "voie 7 chaufferette CM";
END_REGION

REGION Network 34 (STL): spare - CM chan 8
         A     "Epics_to_PLC"."spare-CM-8".cmdSet;
         S     "voie 8 chaufferette CM";
         A     "Epics_to_PLC"."spare-CM-8".cmdRst;
         R     "voie 8 chaufferette CM";
END_REGION

REGION Network 35 (STL): spare - CM chan 10
         A     "Epics_to_PLC"."spare-CM-10".cmdSet;
         S     "voie 10 chaufferette CM";
         A     "Epics_to_PLC"."spare-CM-10".cmdRst;
         R     "voie 10 chaufferette CM";
END_REGION

REGION Network 36 (STL): spare - CM chan 12
         A     "Epics_to_PLC"."spare-CM-12".cmdSet;
         S     "voie 12 chaufferette CM";
         A     "Epics_to_PLC"."spare-CM-12".cmdRst;
         R     "voie 12 chaufferette CM";
END_REGION

REGION Network 37 (STL): Bit commands
         A     "Epics_to_PLC".cmdAutoMode;
         R     "Graph/manuelle";
         A     "Epics_to_PLC".cmdManMode;
         S     "Graph/manuelle";
         A     "Epics_to_PLC".cmdGrafcetInit;
         =     "MettreEtatInitial";
         A     "Epics_to_PLC".cmdGrafcetErrRst;
         =     "AcquitterErreurGraph";
         A     "Epics_to_PLC".cmdStartConditioning;
         =     "CmdVanneEtatCdt";
         A     "Epics_to_PLC".cmdCondOK;
         =     "CdtInfraOk";
         A     "Epics_to_PLC".cmdCondERR;
         =     "CdtInfraErreur";
         A     "Epics_to_PLC".cmdStartLN2cooling;
         =     "DmdMefAzote";
         A     "Epics_to_PLC".cmdStartLHecooling;
         =     "DmdMefHelium";
         A     "Epics_to_PLC".cmdStart2Kmode;
         =     "DmdMode2K";
         A     "Epics_to_PLC".cmdStop2Kmode;
         =     "DmdArretMode2k";
         A     "Epics_to_PLC".cmdStartSTBYmode;
         =     "DmdModeStandby";
         A     "Epics_to_PLC".cmdStopSTBYmode;
         =     "DmdArretModeStandby";
         A     "Epics_to_PLC".cmdStartHeating;
         =     "StartHeating";
         A     "Epics_to_PLC".cmdStopHeating;
         =     "StopHeating";
END_REGION

REGION Network 38: Real parameters (LHe level PIDs settings)
   RUNG wire#powerrail
      Contact( "Epics_to_PLC".TrigPID_CV01.cmdSet )
      { S7_GenerateENO := "TRUE" } Move(in := "Epics_to_PLC".TrigPID_CV01.cSetV, out1 => "TriggerPIDcv01")
      { S7_GenerateENO := "TRUE" } Move(in := "Epics_to_PLC".TrigPID_CV01.cSetV, out1 => "S8_parameters".TrigPID_CV01)
      R_Coil( "Epics_to_PLC".TrigPID_CV01.cmdSet )
   END_RUNG
   // the same network as SCL:
   // ENO of a box is taken as its EN; it also drops when the box reports an error
   IF "Epics_to_PLC".TrigPID_CV01.cmdSet THEN
       "TriggerPIDcv01" := "Epics_to_PLC".TrigPID_CV01.cSetV;
       "S8_parameters".TrigPID_CV01 := "Epics_to_PLC".TrigPID_CV01.cSetV;
       "Epics_to_PLC".TrigPID_CV01.cmdSet := FALSE;
   END_IF;
END_REGION

